REGION Network 3: Init message
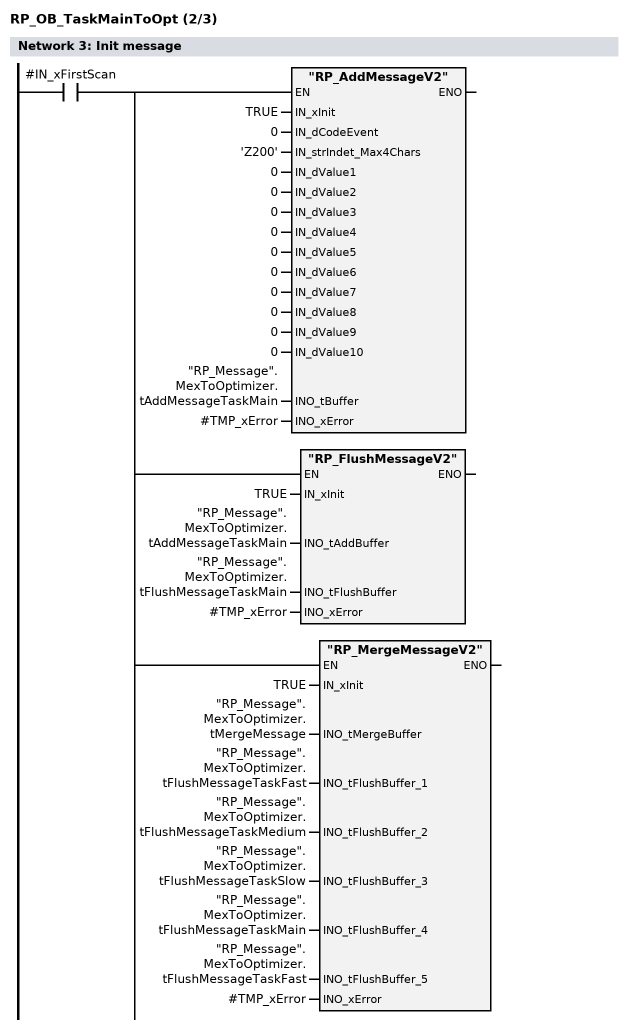
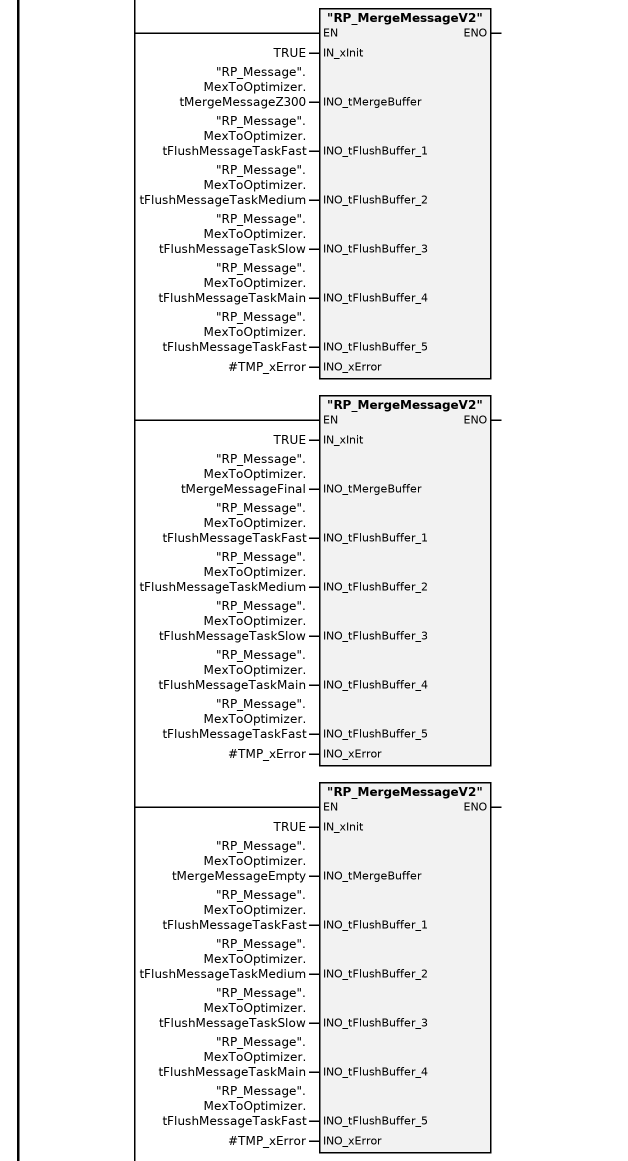
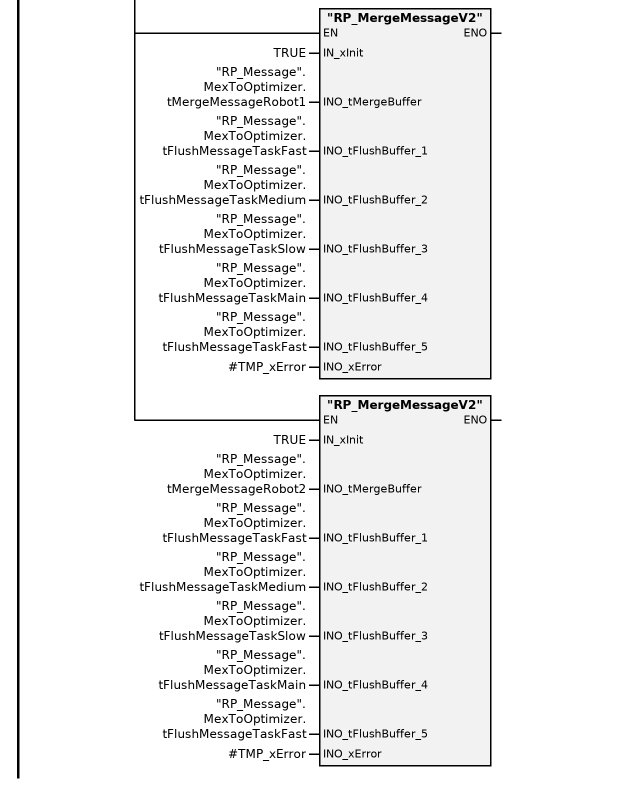
   RUNG wire#powerrail
      Contact( #IN_xFirstScan )
      wire#w1
      "RP_AddMessageV2"(IN_xInit := TRUE, IN_dCodeEvent := 0, IN_strIndet_Max4Chars := 'Z200', IN_dValue1 := 0, IN_dValue2 := 0, IN_dValue3 := 0, IN_dValue4 := 0, IN_dValue5 := 0, IN_dValue6 := 0, IN_dValue7 := 0, IN_dValue8 := 0, IN_dValue9 := 0, IN_dValue10 := 0, INO_tBuffer := "RP_Message".MexToOptimizer.tAddMessageTaskMain, INO_xError := #TMP_xError)
   END_RUNG
   RUNG wire#w1
      "RP_FlushMessageV2"(IN_xInit := TRUE, INO_tAddBuffer := "RP_Message".MexToOptimizer.tAddMessageTaskMain, INO_tFlushBuffer := "RP_Message".MexToOptimizer.tFlushMessageTaskMain, INO_xError := #TMP_xError)
   END_RUNG
   RUNG wire#w1
      "RP_MergeMessageV2"(IN_xInit := TRUE, INO_tMergeBuffer := "RP_Message".MexToOptimizer.tMergeMessage, INO_tFlushBuffer_1 := "RP_Message".MexToOptimizer.tFlushMessageTaskFast, INO_tFlushBuffer_2 := "RP_Message".MexToOptimizer.tFlushMessageTaskMedium, INO_tFlushBuffer_3 := "RP_Message".MexToOptimizer.tFlushMessageTaskSlow, INO_tFlushBuffer_4 := "RP_Message".MexToOptimizer.tFlushMessageTaskMain, INO_tFlushBuffer_5 := "RP_Message".MexToOptimizer.tFlushMessageTaskFast, INO_xError := #TMP_xError)
   END_RUNG
   RUNG wire#w1
      "RP_MergeMessageV2"(IN_xInit := TRUE, INO_tMergeBuffer := "RP_Message".MexToOptimizer.tMergeMessageZ300, INO_tFlushBuffer_1 := "RP_Message".MexToOptimizer.tFlushMessageTaskFast, INO_tFlushBuffer_2 := "RP_Message".MexToOptimizer.tFlushMessageTaskMedium, INO_tFlushBuffer_3 := "RP_Message".MexToOptimizer.tFlushMessageTaskSlow, INO_tFlushBuffer_4 := "RP_Message".MexToOptimizer.tFlushMessageTaskMain, INO_tFlushBuffer_5 := "RP_Message".MexToOptimizer.tFlushMessageTaskFast, INO_xError := #TMP_xError)
   END_RUNG
   RUNG wire#w1
      "RP_MergeMessageV2"(IN_xInit := TRUE, INO_tMergeBuffer := "RP_Message".MexToOptimizer.tMergeMessageFinal, INO_tFlushBuffer_1 := "RP_Message".MexToOptimizer.tFlushMessageTaskFast, INO_tFlushBuffer_2 := "RP_Message".MexToOptimizer.tFlushMessageTaskMedium, INO_tFlushBuffer_3 := "RP_Message".MexToOptimizer.tFlushMessageTaskSlow, INO_tFlushBuffer_4 := "RP_Message".MexToOptimizer.tFlushMessageTaskMain, INO_tFlushBuffer_5 := "RP_Message".MexToOptimizer.tFlushMessageTaskFast, INO_xError := #TMP_xError)
   END_RUNG
   RUNG wire#w1
      "RP_MergeMessageV2"(IN_xInit := TRUE, INO_tMergeBuffer := "RP_Message".MexToOptimizer.tMergeMessageEmpty, INO_tFlushBuffer_1 := "RP_Message".MexToOptimizer.tFlushMessageTaskFast, INO_tFlushBuffer_2 := "RP_Message".MexToOptimizer.tFlushMessageTaskMedium, INO_tFlushBuffer_3 := "RP_Message".MexToOptimizer.tFlushMessageTaskSlow, INO_tFlushBuffer_4 := "RP_Message".MexToOptimizer.tFlushMessageTaskMain, INO_tFlushBuffer_5 := "RP_Message".MexToOptimizer.tFlushMessageTaskFast, INO_xError := #TMP_xError)
   END_RUNG
   RUNG wire#w1
      "RP_MergeMessageV2"(IN_xInit := TRUE, INO_tMergeBuffer := "RP_Message".MexToOptimizer.tMergeMessageRobot1, INO_tFlushBuffer_1 := "RP_Message".MexToOptimizer.tFlushMessageTaskFast, INO_tFlushBuffer_2 := "RP_Message".MexToOptimizer.tFlushMessageTaskMedium, INO_tFlushBuffer_3 := "RP_Message".MexToOptimizer.tFlushMessageTaskSlow, INO_tFlushBuffer_4 := "RP_Message".MexToOptimizer.tFlushMessageTaskMain, INO_tFlushBuffer_5 := "RP_Message".MexToOptimizer.tFlushMessageTaskFast, INO_xError := #TMP_xError)
   END_RUNG
   RUNG wire#w1
      "RP_MergeMessageV2"(IN_xInit := TRUE, INO_tMergeBuffer := "RP_Message".MexToOptimizer.tMergeMessageRobot2, INO_tFlushBuffer_1 := "RP_Message".MexToOptimizer.tFlushMessageTaskFast, INO_tFlushBuffer_2 := "RP_Message".MexToOptimizer.tFlushMessageTaskMedium, INO_tFlushBuffer_3 := "RP_Message".MexToOptimizer.tFlushMessageTaskSlow, INO_tFlushBuffer_4 := "RP_Message".MexToOptimizer.tFlushMessageTaskMain, INO_tFlushBuffer_5 := "RP_Message".MexToOptimizer.tFlushMessageTaskFast, INO_xError := #TMP_xError)
   END_RUNG
   // the same network as SCL:
   IF #IN_xFirstScan THEN
       "RP_AddMessageV2"(IN_xInit := TRUE,
                         IN_dCodeEvent := 0,
                         IN_strIndet_Max4Chars := 'Z200',
                         IN_dValue1 := 0,
                         IN_dValue2 := 0,
                         IN_dValue3 := 0,
                         IN_dValue4 := 0,
                         IN_dValue5 := 0,
                         IN_dValue6 := 0,
                         IN_dValue7 := 0,
                         IN_dValue8 := 0,
                         IN_dValue9 := 0,
                         IN_dValue10 := 0,
                         INO_tBuffer := "RP_Message".MexToOptimizer.tAddMessageTaskMain,
                         INO_xError := #TMP_xError);
       "RP_FlushMessageV2"(IN_xInit := TRUE,
                           INO_tAddBuffer := "RP_Message".MexToOptimizer.tAddMessageTaskMain,
                           INO_tFlushBuffer := "RP_Message".MexToOptimizer.tFlushMessageTaskMain,
                           INO_xError := #TMP_xError);
       "RP_MergeMessageV2"(IN_xInit := TRUE,
                           INO_tMergeBuffer := "RP_Message".MexToOptimizer.tMergeMessage,
                           INO_tFlushBuffer_1 := "RP_Message".MexToOptimizer.tFlushMessageTaskFast,
                           INO_tFlushBuffer_2 := "RP_Message".MexToOptimizer.tFlushMessageTaskMedium,
                           INO_tFlushBuffer_3 := "RP_Message".MexToOptimizer.tFlushMessageTaskSlow,
                           INO_tFlushBuffer_4 := "RP_Message".MexToOptimizer.tFlushMessageTaskMain,
                           INO_tFlushBuffer_5 := "RP_Message".MexToOptimizer.tFlushMessageTaskFast,
                           INO_xError := #TMP_xError);
       "RP_MergeMessageV2"(IN_xInit := TRUE,
                           INO_tMergeBuffer := "RP_Message".MexToOptimizer.tMergeMessageZ300,
                           INO_tFlushBuffer_1 := "RP_Message".MexToOptimizer.tFlushMessageTaskFast,
                           INO_tFlushBuffer_2 := "RP_Message".MexToOptimizer.tFlushMessageTaskMedium,
                           INO_tFlushBuffer_3 := "RP_Message".MexToOptimizer.tFlushMessageTaskSlow,
                           INO_tFlushBuffer_4 := "RP_Message".MexToOptimizer.tFlushMessageTaskMain,
                           INO_tFlushBuffer_5 := "RP_Message".MexToOptimizer.tFlushMessageTaskFast,
                           INO_xError := #TMP_xError);
       "RP_MergeMessageV2"(IN_xInit := TRUE,
                           INO_tMergeBuffer := "RP_Message".MexToOptimizer.tMergeMessageFinal,
                           INO_tFlushBuffer_1 := "RP_Message".MexToOptimizer.tFlushMessageTaskFast,
                           INO_tFlushBuffer_2 := "RP_Message".MexToOptimizer.tFlushMessageTaskMedium,
                           INO_tFlushBuffer_3 := "RP_Message".MexToOptimizer.tFlushMessageTaskSlow,
                           INO_tFlushBuffer_4 := "RP_Message".MexToOptimizer.tFlushMessageTaskMain,
                           INO_tFlushBuffer_5 := "RP_Message".MexToOptimizer.tFlushMessageTaskFast,
                           INO_xError := #TMP_xError);
       "RP_MergeMessageV2"(IN_xInit := TRUE,
                           INO_tMergeBuffer := "RP_Message".MexToOptimizer.tMergeMessageEmpty,
                           INO_tFlushBuffer_1 := "RP_Message".MexToOptimizer.tFlushMessageTaskFast,
                           INO_tFlushBuffer_2 := "RP_Message".MexToOptimizer.tFlushMessageTaskMedium,
                           INO_tFlushBuffer_3 := "RP_Message".MexToOptimizer.tFlushMessageTaskSlow,
                           INO_tFlushBuffer_4 := "RP_Message".MexToOptimizer.tFlushMessageTaskMain,
                           INO_tFlushBuffer_5 := "RP_Message".MexToOptimizer.tFlushMessageTaskFast,
                           INO_xError := #TMP_xError);
       "RP_MergeMessageV2"(IN_xInit := TRUE,
                           INO_tMergeBuffer := "RP_Message".MexToOptimizer.tMergeMessageRobot1,
                           INO_tFlushBuffer_1 := "RP_Message".MexToOptimizer.tFlushMessageTaskFast,
                           INO_tFlushBuffer_2 := "RP_Message".MexToOptimizer.tFlushMessageTaskMedium,
                           INO_tFlushBuffer_3 := "RP_Message".MexToOptimizer.tFlushMessageTaskSlow,
                           INO_tFlushBuffer_4 := "RP_Message".MexToOptimizer.tFlushMessageTaskMain,
                           INO_tFlushBuffer_5 := "RP_Message".MexToOptimizer.tFlushMessageTaskFast,
                           INO_xError := #TMP_xError);
       "RP_MergeMessageV2"(IN_xInit := TRUE,
                           INO_tMergeBuffer := "RP_Message".MexToOptimizer.tMergeMessageRobot2,
                           INO_tFlushBuffer_1 := "RP_Message".MexToOptimizer.tFlushMessageTaskFast,
                           INO_tFlushBuffer_2 := "RP_Message".MexToOptimizer.tFlushMessageTaskMedium,
                           INO_tFlushBuffer_3 := "RP_Message".MexToOptimizer.tFlushMessageTaskSlow,
                           INO_tFlushBuffer_4 := "RP_Message".MexToOptimizer.tFlushMessageTaskMain,
                           INO_tFlushBuffer_5 := "RP_Message".MexToOptimizer.tFlushMessageTaskFast,
                           INO_xError := #TMP_xError);
   END_IF;
END_REGION

REGION Network 4: Flush message
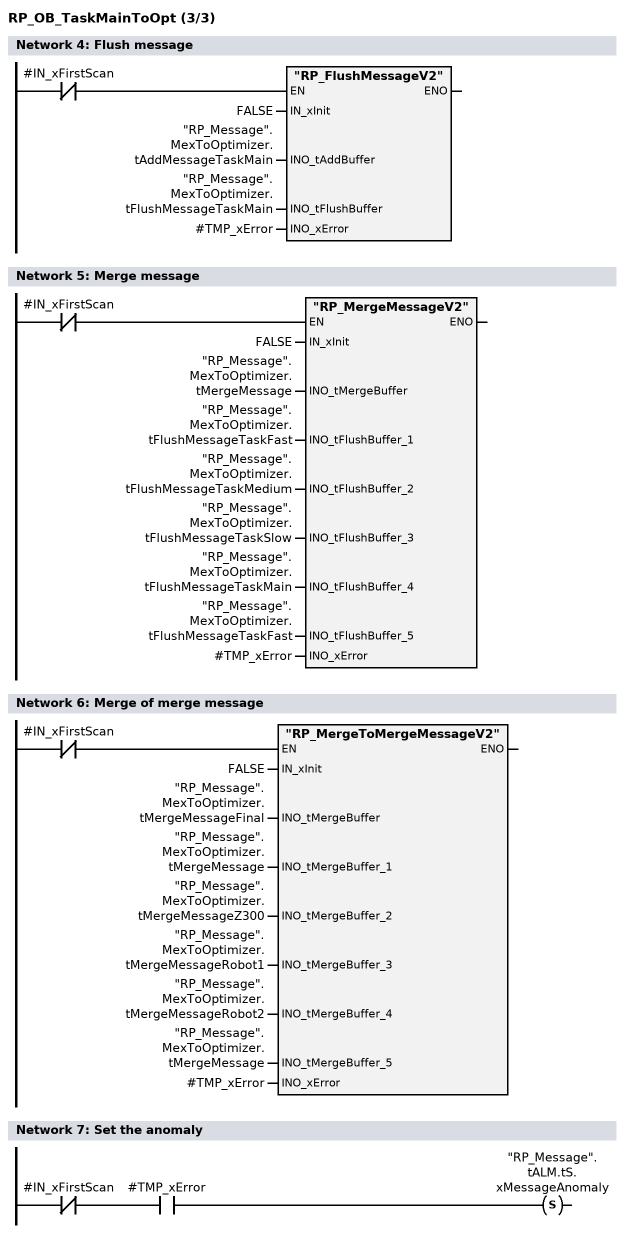
   RUNG wire#powerrail
      I_Contact( #IN_xFirstScan )
      "RP_FlushMessageV2"(IN_xInit := FALSE, INO_tAddBuffer := "RP_Message".MexToOptimizer.tAddMessageTaskMain, INO_tFlushBuffer := "RP_Message".MexToOptimizer.tFlushMessageTaskMain, INO_xError := #TMP_xError)
   END_RUNG
   // the same network as SCL:
   IF NOT #IN_xFirstScan THEN
       "RP_FlushMessageV2"(IN_xInit := FALSE,
                           INO_tAddBuffer := "RP_Message".MexToOptimizer.tAddMessageTaskMain,
                           INO_tFlushBuffer := "RP_Message".MexToOptimizer.tFlushMessageTaskMain,
                           INO_xError := #TMP_xError);
   END_IF;
END_REGION

REGION Network 5: Merge message
   RUNG wire#powerrail
      I_Contact( #IN_xFirstScan )
      "RP_MergeMessageV2"(IN_xInit := FALSE, INO_tMergeBuffer := "RP_Message".MexToOptimizer.tMergeMessage, INO_tFlushBuffer_1 := "RP_Message".MexToOptimizer.tFlushMessageTaskFast, INO_tFlushBuffer_2 := "RP_Message".MexToOptimizer.tFlushMessageTaskMedium, INO_tFlushBuffer_3 := "RP_Message".MexToOptimizer.tFlushMessageTaskSlow, INO_tFlushBuffer_4 := "RP_Message".MexToOptimizer.tFlushMessageTaskMain, INO_tFlushBuffer_5 := "RP_Message".MexToOptimizer.tFlushMessageTaskFast, INO_xError := #TMP_xError)
   END_RUNG
   // the same network as SCL:
   IF NOT #IN_xFirstScan THEN
       "RP_MergeMessageV2"(IN_xInit := FALSE,
                           INO_tMergeBuffer := "RP_Message".MexToOptimizer.tMergeMessage,
                           INO_tFlushBuffer_1 := "RP_Message".MexToOptimizer.tFlushMessageTaskFast,
                           INO_tFlushBuffer_2 := "RP_Message".MexToOptimizer.tFlushMessageTaskMedium,
                           INO_tFlushBuffer_3 := "RP_Message".MexToOptimizer.tFlushMessageTaskSlow,
                           INO_tFlushBuffer_4 := "RP_Message".MexToOptimizer.tFlushMessageTaskMain,
                           INO_tFlushBuffer_5 := "RP_Message".MexToOptimizer.tFlushMessageTaskFast,
                           INO_xError := #TMP_xError);
   END_IF;
END_REGION

REGION Network 6: Merge of merge message
   RUNG wire#powerrail
      I_Contact( #IN_xFirstScan )
      "RP_MergeToMergeMessageV2"(IN_xInit := FALSE, INO_tMergeBuffer := "RP_Message".MexToOptimizer.tMergeMessageFinal, INO_tMergeBuffer_1 := "RP_Message".MexToOptimizer.tMergeMessage, INO_tMergeBuffer_2 := "RP_Message".MexToOptimizer.tMergeMessageZ300, INO_tMergeBuffer_3 := "RP_Message".MexToOptimizer.tMergeMessageRobot1, INO_tMergeBuffer_4 := "RP_Message".MexToOptimizer.tMergeMessageRobot2, INO_tMergeBuffer_5 := "RP_Message".MexToOptimizer.tMergeMessage, INO_xError := #TMP_xError)
   END_RUNG
   // the same network as SCL:
   IF NOT #IN_xFirstScan THEN
       "RP_MergeToMergeMessageV2"(IN_xInit := FALSE,
                               INO_tMergeBuffer := "RP_Message".MexToOptimizer.tMergeMessageFinal,
                               INO_tMergeBuffer_1 := "RP_Message".MexToOptimizer.tMergeMessage,
                               INO_tMergeBuffer_2 := "RP_Message".MexToOptimizer.tMergeMessageZ300,
                               INO_tMergeBuffer_3 := "RP_Message".MexToOptimizer.tMergeMessageRobot1,
                               INO_tMergeBuffer_4 := "RP_Message".MexToOptimizer.tMergeMessageRobot2,
                               INO_tMergeBuffer_5 := "RP_Message".MexToOptimizer.tMergeMessage,
                               INO_xError := #TMP_xError);
   END_IF;
END_REGION

REGION Network 7: Set the anomaly
   RUNG wire#powerrail
      I_Contact( #IN_xFirstScan )
      Contact( #TMP_xError )
      S_Coil( "RP_Message".tALM.tS.xMessageAnomaly )
   END_RUNG
   // the same network as SCL:
   IF NOT #IN_xFirstScan AND #TMP_xError THEN "RP_Message".tALM.tS.xMessageAnomaly := TRUE; END_IF;
END_REGION

REGION Network 8 (SCL): Moving data to tank
   IF "RP_Message".MexToOptimizer.tMergeMessageFinal.dNumOfMessage > 0 AND
       "RP_Message".MexToOptimizer.tMergeMessageFinal.xInitialized THEN  

       IF  ("RP_Message".MexToOptimizer.tMergeMessageFinal.dNumOfMessage + "RP_Message".tTankMessageForOpt.dNumberOfMessage) < "DMAXNUMMESSAGETANK" THEN
           //Copy the messages on tank
           #TMP_iRet :=  MOVE_BLK_VARIANT(SRC:="RP_Message".MexToOptimizer.tMergeMessageFinal.rgtMessages, 
                           COUNT:=DINT_TO_UDINT("RP_Message".MexToOptimizer.tMergeMessageFinal.dNumOfMessage), 
                           SRC_INDEX:=0, DEST_INDEX:="RP_Message".tTankMessageForOpt.dNumberOfMessage, 
                           DEST=>"RP_Message".tTankMessageForOpt.rgtMessages);

           "RP_Message".tTankMessageForOpt.dNumberOfMessage += "RP_Message".MexToOptimizer.tMergeMessageFinal.dNumOfMessage;
       ELSE
           "RP_Message".tALM.tS.xOptTankFull := TRUE;
       END_IF;

       IF  ("RP_Message".MexToOptimizer.tMergeMessageFinal.dNumOfMessage + "RP_Message".tTankMessageForReport.dNumberOfMessage) < "DMAXNUMMESSAGETANK" THEN
           //Copy the messages on tank
           #TMP_iRet :=  MOVE_BLK_VARIANT(SRC:="RP_Message".MexToOptimizer.tMergeMessageFinal.rgtMessages, 
                           COUNT:=DINT_TO_UDINT("RP_Message".MexToOptimizer.tMergeMessageFinal.dNumOfMessage), 
                           SRC_INDEX:=0, DEST_INDEX:="RP_Message".tTankMessageForReport.dNumberOfMessage, 
                           DEST=>"RP_Message".tTankMessageForReport.rgtMessages);

           "RP_Message".tTankMessageForReport.dNumberOfMessage += "RP_Message".MexToOptimizer.tMergeMessageFinal.dNumOfMessage;
       ELSE
           "RP_Message".tALM.tS.xReportTankFull := TRUE;
       END_IF;

       "RP_Message".MexToOptimizer.tMergeMessageFinal := "RP_Message".MexToOptimizer.tMergeMessageEmpty;

   END_IF;
END_REGION
END_FUNCTION

FUNCTION "RP_OB_TaskFastFromOpt" : Void   // FC20, LAD
{ S7_Optimized_Access := 'TRUE' }
VERSION : 0.1
   VAR_INPUT
      IN_xFirstScan : Bool;
   END_VAR
   VAR_TEMP
      TMP_xError : Bool;
   END_VAR
BEGIN

REGION Network 1
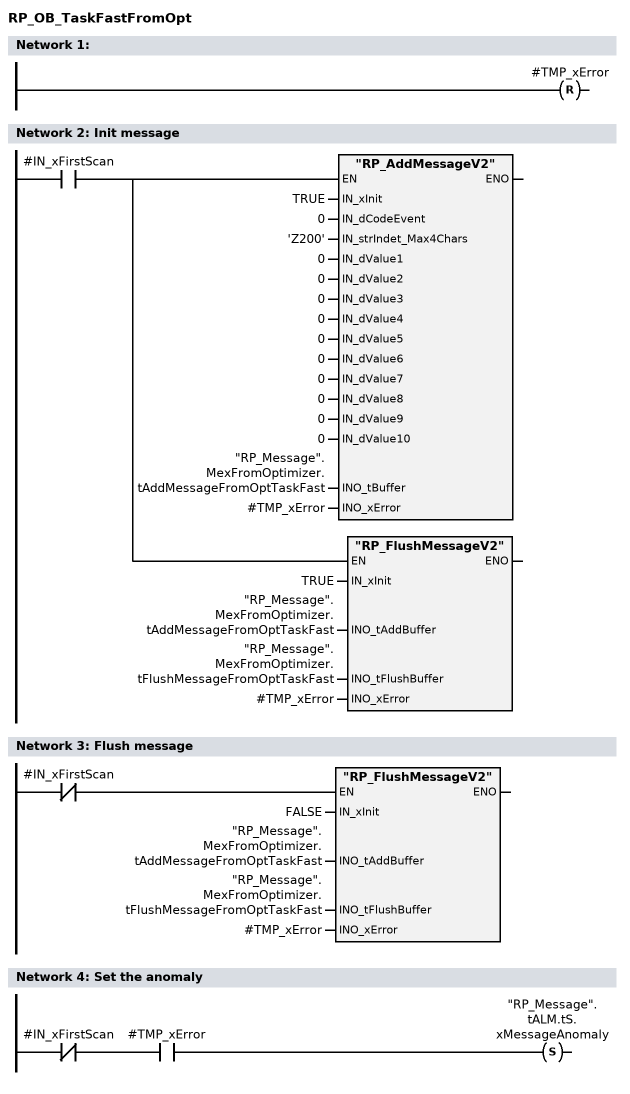
   RUNG wire#powerrail
      R_Coil( #TMP_xError )
   END_RUNG
   // the same network as SCL:
   #TMP_xError := FALSE;
END_REGION

REGION Network 2: Init message
   RUNG wire#powerrail
      Contact( #IN_xFirstScan )
      wire#w1
      "RP_AddMessageV2"(IN_xInit := TRUE, IN_dCodeEvent := 0, IN_strIndet_Max4Chars := 'Z200', IN_dValue1 := 0, IN_dValue2 := 0, IN_dValue3 := 0, IN_dValue4 := 0, IN_dValue5 := 0, IN_dValue6 := 0, IN_dValue7 := 0, IN_dValue8 := 0, IN_dValue9 := 0, IN_dValue10 := 0, INO_tBuffer := "RP_Message".MexFromOptimizer.tAddMessageFromOptTaskFast, INO_xError := #TMP_xError)
   END_RUNG
   RUNG wire#w1
      "RP_FlushMessageV2"(IN_xInit := TRUE, INO_tAddBuffer := "RP_Message".MexFromOptimizer.tAddMessageFromOptTaskFast, INO_tFlushBuffer := "RP_Message".MexFromOptimizer.tFlushMessageFromOptTaskFast, INO_xError := #TMP_xError)
   END_RUNG
   // the same network as SCL:
   IF #IN_xFirstScan THEN
       "RP_AddMessageV2"(IN_xInit := TRUE,
                         IN_dCodeEvent := 0,
                         IN_strIndet_Max4Chars := 'Z200',
                         IN_dValue1 := 0,
                         IN_dValue2 := 0,
                         IN_dValue3 := 0,
                         IN_dValue4 := 0,
                         IN_dValue5 := 0,
                         IN_dValue6 := 0,
                         IN_dValue7 := 0,
                         IN_dValue8 := 0,
                         IN_dValue9 := 0,
                         IN_dValue10 := 0,
                         INO_tBuffer := "RP_Message".MexFromOptimizer.tAddMessageFromOptTaskFast,
                         INO_xError := #TMP_xError);
       "RP_FlushMessageV2"(IN_xInit := TRUE,
                           INO_tAddBuffer := "RP_Message".MexFromOptimizer.tAddMessageFromOptTaskFast,
                           INO_tFlushBuffer := "RP_Message".MexFromOptimizer.tFlushMessageFromOptTaskFast,
                           INO_xError := #TMP_xError);
   END_IF;
END_REGION

REGION Network 3: Flush message
   RUNG wire#powerrail
      I_Contact( #IN_xFirstScan )
      "RP_FlushMessageV2"(IN_xInit := FALSE, INO_tAddBuffer := "RP_Message".MexFromOptimizer.tAddMessageFromOptTaskFast, INO_tFlushBuffer := "RP_Message".MexFromOptimizer.tFlushMessageFromOptTaskFast, INO_xError := #TMP_xError)
   END_RUNG
   // the same network as SCL:
   IF NOT #IN_xFirstScan THEN
       "RP_FlushMessageV2"(IN_xInit := FALSE,
                           INO_tAddBuffer := "RP_Message".MexFromOptimizer.tAddMessageFromOptTaskFast,
                           INO_tFlushBuffer := "RP_Message".MexFromOptimizer.tFlushMessageFromOptTaskFast,
                           INO_xError := #TMP_xError);
   END_IF;
END_REGION

REGION Network 4: Set the anomaly
   RUNG wire#powerrail
      I_Contact( #IN_xFirstScan )
      Contact( #TMP_xError )
      S_Coil( "RP_Message".tALM.tS.xMessageAnomaly )
   END_RUNG
   // the same network as SCL:
   IF NOT #IN_xFirstScan AND #TMP_xError THEN "RP_Message".tALM.tS.xMessageAnomaly := TRUE; END_IF;
END_REGION
END_FUNCTION

FUNCTION "RP_OB_TaskSlowFromOpt" : Void   // FC21, LAD
{ S7_Optimized_Access := 'TRUE' }
VERSION : 0.1
   VAR_INPUT
      IN_xFirstScan : Bool;
   END_VAR
   VAR_TEMP
      TMP_xError : Bool;
   END_VAR
BEGIN

REGION Network 1
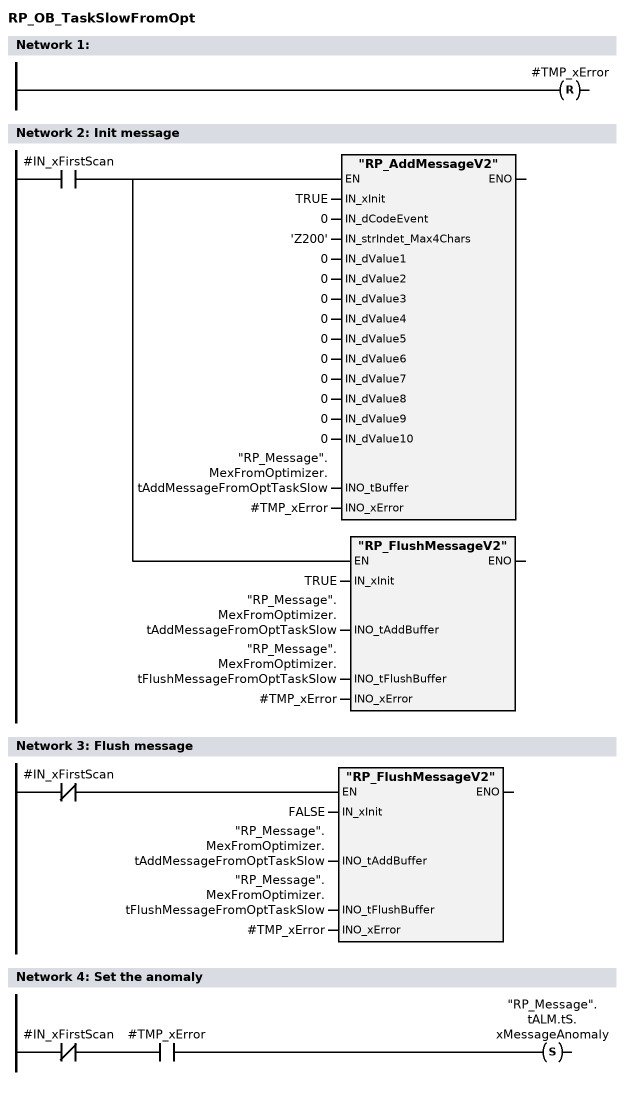
   RUNG wire#powerrail
      R_Coil( #TMP_xError )
   END_RUNG
   // the same network as SCL:
   #TMP_xError := FALSE;
END_REGION

REGION Network 2: Init message
   RUNG wire#powerrail
      Contact( #IN_xFirstScan )
      wire#w1
      "RP_AddMessageV2"(IN_xInit := TRUE, IN_dCodeEvent := 0, IN_strIndet_Max4Chars := 'Z200', IN_dValue1 := 0, IN_dValue2 := 0, IN_dValue3 := 0, IN_dValue4 := 0, IN_dValue5 := 0, IN_dValue6 := 0, IN_dValue7 := 0, IN_dValue8 := 0, IN_dValue9 := 0, IN_dValue10 := 0, INO_tBuffer := "RP_Message".MexFromOptimizer.tAddMessageFromOptTaskSlow, INO_xError := #TMP_xError)
   END_RUNG
   RUNG wire#w1
      "RP_FlushMessageV2"(IN_xInit := TRUE, INO_tAddBuffer := "RP_Message".MexFromOptimizer.tAddMessageFromOptTaskSlow, INO_tFlushBuffer := "RP_Message".MexFromOptimizer.tFlushMessageFromOptTaskSlow, INO_xError := #TMP_xError)
   END_RUNG
   // the same network as SCL:
   IF #IN_xFirstScan THEN
       "RP_AddMessageV2"(IN_xInit := TRUE,
                         IN_dCodeEvent := 0,
                         IN_strIndet_Max4Chars := 'Z200',
                         IN_dValue1 := 0,
                         IN_dValue2 := 0,
                         IN_dValue3 := 0,
                         IN_dValue4 := 0,
                         IN_dValue5 := 0,
                         IN_dValue6 := 0,
                         IN_dValue7 := 0,
                         IN_dValue8 := 0,
                         IN_dValue9 := 0,
                         IN_dValue10 := 0,
                         INO_tBuffer := "RP_Message".MexFromOptimizer.tAddMessageFromOptTaskSlow,
                         INO_xError := #TMP_xError);
       "RP_FlushMessageV2"(IN_xInit := TRUE,
                           INO_tAddBuffer := "RP_Message".MexFromOptimizer.tAddMessageFromOptTaskSlow,
                           INO_tFlushBuffer := "RP_Message".MexFromOptimizer.tFlushMessageFromOptTaskSlow,
                           INO_xError := #TMP_xError);
   END_IF;
END_REGION

REGION Network 3: Flush message
   RUNG wire#powerrail
      I_Contact( #IN_xFirstScan )
      "RP_FlushMessageV2"(IN_xInit := FALSE, INO_tAddBuffer := "RP_Message".MexFromOptimizer.tAddMessageFromOptTaskSlow, INO_tFlushBuffer := "RP_Message".MexFromOptimizer.tFlushMessageFromOptTaskSlow, INO_xError := #TMP_xError)
   END_RUNG
   // the same network as SCL:
   IF NOT #IN_xFirstScan THEN
       "RP_FlushMessageV2"(IN_xInit := FALSE,
                           INO_tAddBuffer := "RP_Message".MexFromOptimizer.tAddMessageFromOptTaskSlow,
                           INO_tFlushBuffer := "RP_Message".MexFromOptimizer.tFlushMessageFromOptTaskSlow,
                           INO_xError := #TMP_xError);
   END_IF;
END_REGION

REGION Network 4: Set the anomaly
   RUNG wire#powerrail
      I_Contact( #IN_xFirstScan )
      Contact( #TMP_xError )
      S_Coil( "RP_Message".tALM.tS.xMessageAnomaly )
   END_RUNG
   // the same network as SCL:
   IF NOT #IN_xFirstScan AND #TMP_xError THEN "RP_Message".tALM.tS.xMessageAnomaly := TRUE; END_IF;
END_REGION
END_FUNCTION

FUNCTION "RP_OB_TaskMainFromOpt" : Void   // FC22, LAD
{ S7_Optimized_Access := 'TRUE' }
VERSION : 0.1
   VAR_INPUT
      IN_xFirstScan : Bool;
   END_VAR
   VAR_TEMP
      TMP_xError : Bool;
      TMP_iRet : Int;
      TMP_dwValue : DWord;
   END_VAR
BEGIN

REGION Network 1: Reset temporary
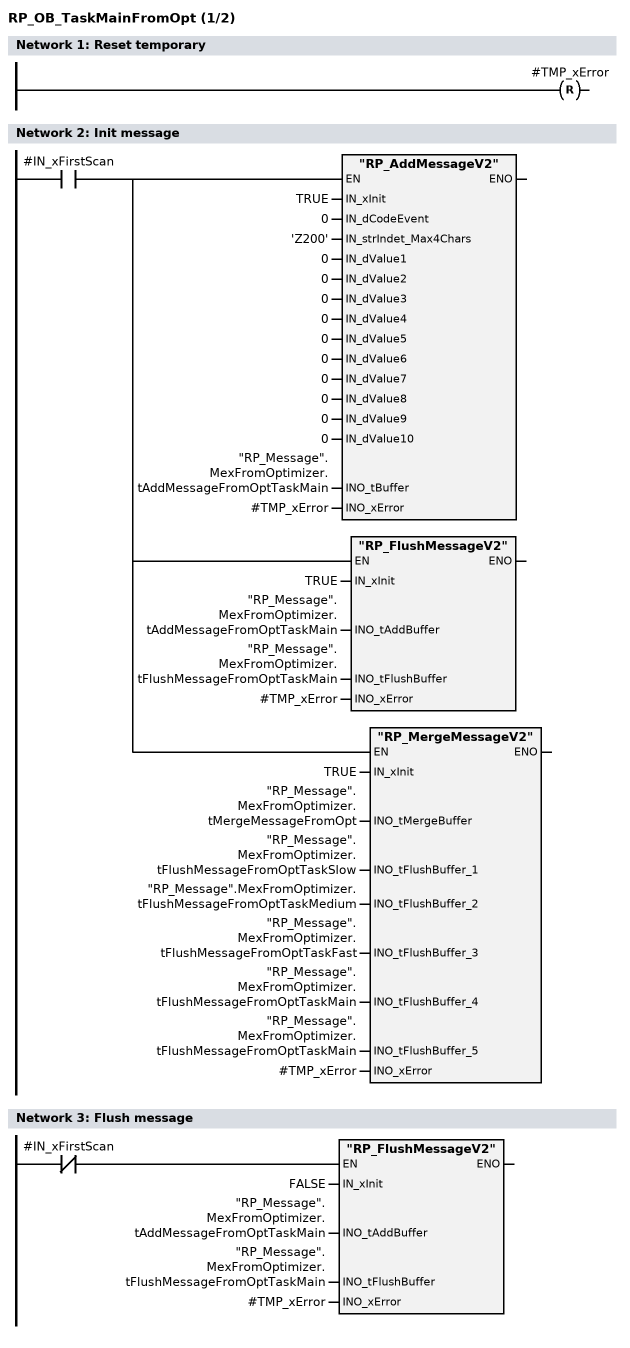
   RUNG wire#powerrail
      R_Coil( #TMP_xError )
   END_RUNG
   // the same network as SCL:
   #TMP_xError := FALSE;
END_REGION

REGION Network 2: Init message
   RUNG wire#powerrail
      Contact( #IN_xFirstScan )
      wire#w1
      "RP_AddMessageV2"(IN_xInit := TRUE, IN_dCodeEvent := 0, IN_strIndet_Max4Chars := 'Z200', IN_dValue1 := 0, IN_dValue2 := 0, IN_dValue3 := 0, IN_dValue4 := 0, IN_dValue5 := 0, IN_dValue6 := 0, IN_dValue7 := 0, IN_dValue8 := 0, IN_dValue9 := 0, IN_dValue10 := 0, INO_tBuffer := "RP_Message".MexFromOptimizer.tAddMessageFromOptTaskMain, INO_xError := #TMP_xError)
   END_RUNG
   RUNG wire#w1
      "RP_FlushMessageV2"(IN_xInit := TRUE, INO_tAddBuffer := "RP_Message".MexFromOptimizer.tAddMessageFromOptTaskMain, INO_tFlushBuffer := "RP_Message".MexFromOptimizer.tFlushMessageFromOptTaskMain, INO_xError := #TMP_xError)
   END_RUNG
   RUNG wire#w1
      "RP_MergeMessageV2"(IN_xInit := TRUE, INO_tMergeBuffer := "RP_Message".MexFromOptimizer.tMergeMessageFromOpt, INO_tFlushBuffer_1 := "RP_Message".MexFromOptimizer.tFlushMessageFromOptTaskSlow, INO_tFlushBuffer_2 := "RP_Message".MexFromOptimizer.tFlushMessageFromOptTaskMedium, INO_tFlushBuffer_3 := "RP_Message".MexFromOptimizer.tFlushMessageFromOptTaskFast, INO_tFlushBuffer_4 := "RP_Message".MexFromOptimizer.tFlushMessageFromOptTaskMain, INO_tFlushBuffer_5 := "RP_Message".MexFromOptimizer.tFlushMessageFromOptTaskMain, INO_xError := #TMP_xError)
   END_RUNG
   // the same network as SCL:
   IF #IN_xFirstScan THEN
       "RP_AddMessageV2"(IN_xInit := TRUE,
                         IN_dCodeEvent := 0,
                         IN_strIndet_Max4Chars := 'Z200',
                         IN_dValue1 := 0,
                         IN_dValue2 := 0,
                         IN_dValue3 := 0,
                         IN_dValue4 := 0,
                         IN_dValue5 := 0,
                         IN_dValue6 := 0,
                         IN_dValue7 := 0,
                         IN_dValue8 := 0,
                         IN_dValue9 := 0,
                         IN_dValue10 := 0,
                         INO_tBuffer := "RP_Message".MexFromOptimizer.tAddMessageFromOptTaskMain,
                         INO_xError := #TMP_xError);
       "RP_FlushMessageV2"(IN_xInit := TRUE,
                           INO_tAddBuffer := "RP_Message".MexFromOptimizer.tAddMessageFromOptTaskMain,
                           INO_tFlushBuffer := "RP_Message".MexFromOptimizer.tFlushMessageFromOptTaskMain,
                           INO_xError := #TMP_xError);
       "RP_MergeMessageV2"(IN_xInit := TRUE,
                           INO_tMergeBuffer := "RP_Message".MexFromOptimizer.tMergeMessageFromOpt,
                           INO_tFlushBuffer_1 := "RP_Message".MexFromOptimizer.tFlushMessageFromOptTaskSlow,
                           INO_tFlushBuffer_2 := "RP_Message".MexFromOptimizer.tFlushMessageFromOptTaskMedium,
                           INO_tFlushBuffer_3 := "RP_Message".MexFromOptimizer.tFlushMessageFromOptTaskFast,
                           INO_tFlushBuffer_4 := "RP_Message".MexFromOptimizer.tFlushMessageFromOptTaskMain,
                           INO_tFlushBuffer_5 := "RP_Message".MexFromOptimizer.tFlushMessageFromOptTaskMain,
                           INO_xError := #TMP_xError);
   END_IF;
END_REGION

REGION Network 3: Flush message
   RUNG wire#powerrail
      I_Contact( #IN_xFirstScan )
      "RP_FlushMessageV2"(IN_xInit := FALSE, INO_tAddBuffer := "RP_Message".MexFromOptimizer.tAddMessageFromOptTaskMain, INO_tFlushBuffer := "RP_Message".MexFromOptimizer.tFlushMessageFromOptTaskMain, INO_xError := #TMP_xError)
   END_RUNG
   // the same network as SCL:
   IF NOT #IN_xFirstScan THEN
       "RP_FlushMessageV2"(IN_xInit := FALSE,
                           INO_tAddBuffer := "RP_Message".MexFromOptimizer.tAddMessageFromOptTaskMain,
                           INO_tFlushBuffer := "RP_Message".MexFromOptimizer.tFlushMessageFromOptTaskMain,
                           INO_xError := #TMP_xError);
   END_IF;
END_REGION

REGION Network 4: Merge message